1030 '~Spare MB2[32].6'; 1031 '~Spare MB2[32].7'; 1032 '~S001R13CN.I.StudWld2Rdy - Robot Stud Weld Controller 2 Not Ready MB2[32].8'; 1033 '~S001R13CN.I.Rvt2RdyToOperate - Robot Rivet Controller 2 Not Ready MB2[32].9'; 1034 '~S001R13CN.Ix.LaserWldOn - Robot Laser In No Cut MB2[32].10'; 1035 '~S001R13CN.Ix.GlassNotPres - Robot Laser Glass Not Present MB2[32].11'; 1036 '~S001R13CN.Ix.LaserHeadRdy - Robot Laser Head Not Ready MB2[32].12'; 1037 '~S001R13CN.Ix.ChillerOn - Robot Laser Chiller Not On MB2[32].13'; 1038 '~S001R13CN.Ix.GasOn - Robot Gas Not On MB2[32].14'; 1039 '~S001R13 Power Meter Not Ready MB2[32].15'; 1040 '~S001R13 No Wire Present Replace Barrel MB2[32].16'; 1041 '~S001R13 Wire Feeder Fault Timer MB2[32].17'; 1042 '~S001R13CN.Ix.NRFlt - Robot Nut Runner Not Ready MB2[32].18'; 1043 '~Spare MB2[32].19'; 1044 '~S001R13CN.M.WrongRivetAtNose - Remove Wrong Rivet At Nose MB2[32].20'; 1045 '~S001R13CN.M.DisableRbtDrvs - In Rivet Zone But Riveter Not In Auto MB2[32].21'; 1046 '~S001R13CN.I.Rvt1SystemInAuto - Rivet Controller 1 Not In Auto MB2[32].22'; 1047 '~S001R13CN.I.Rvt2SystemInAuto - Rivet Controller 2 Not In Auto MB2[32].23'; 1048 '~S001R13CN.M.RvtC1ReelCtr.DN - Reel Change Required MB2[32].24'; 1049 '~S001R13CN.M.RvtC2ReelCtr.DN - Reel Change Required MB2[32].25'; 1050 '~S001R13CN.M.AbortSkipRemain - SkipRemaining Aborted, Reset At Rbt Controller Is Required MB2[32].26'; 1051 '~Spare MB2[32].27'; 1052 '~Spare MB2[32].28'; 1053 '~Spare MB2[32].29'; 1054 '~Spare MB2[32].30'; 1055 '~Spare MB2[32].31'; 1056 '~Spare MB2[33].0'; 1057 '~Spare MB2[33].1'; 1058 '~Spare MB2[33].2'; 1059 '~Spare MB2[33].3'; 1060 '~Spare MB2[33].4'; 1061 '~Spare MB2[33].5'; 1062 '~Spare MB2[33].6'; 1063 '~Spare MB2[33].7'; 1064 '~Spare MB2[33].8'; 1065 '~Spare MB2[33].9'; 1066 '~Spare MB2[33].10'; 1067 '~Spare MB2[33].11'; 1068 '~Spare MB2[33].12'; 1069 '~Spare MB2[33].13'; 1070 '~Spare MB2[33].14'; 1071 '~Spare MB2[33].15'; 1072 '~Spare MB2[33].16'; 1073 '~Spare MB2[33].17'; 1074 '~Spare MB2[33].18'; 1075 '~Spare MB2[33].19'; 1076 '~Spare MB2[33].20'; 1077 '~Spare MB2[33].21'; 1078 '~Spare MB2[33].22'; 1079 '~Spare MB2[33].23'; 1080 '~Spare MB2[33].24'; 1081 '~Spare MB2[33].25'; 1082 '~Spare MB2[33].26'; 1083 '~Spare MB2[33].27'; 1084 '~Spare MB2[33].28'; 1085 '~Spare MB2[33].29'; 1086 '~Spare MB2[33].30'; 1087 '~Spare MB2[33].31'; 1088 '~Spare MB2[34].0'; 1089 '~Spare MB2[34].1'; 1090 '~Spare MB2[34].2'; 1091 '~Spare MB2[34].3'; 1092 '~Spare MB2[34].4'; 1093 '~Spare MB2[34].5'; 1094 '~Spare MB2[34].6'; 1095 '~Spare MB2[34].7'; 1096 '~Spare MB2[34].8'; 1097 '~Spare MB2[34].9'; 1098 '~Spare MB2[34].10'; 1099 '~Spare MB2[34].11'; 1100 '~Spare MB2[34].12'; 1101 '~Spare MB2[34].13'; 1102 '~Spare MB2[34].14'; 1103 '~Spare MB2[34].15'; 1104 '~Spare MB2[34].16'; 1105 '~Spare MB2[34].17'; 1106 '~Spare MB2[34].18'; 1107 '~Spare MB2[34].19'; 1108 '~Spare MB2[34].20'; 1109 '~Spare MB2[34].21'; 1110 '~Spare MB2[34].22'; 1111 '~Spare MB2[34].23'; 1112 '~Spare MB2[34].24'; 1113 '~Spare MB2[34].25'; 1114 '~Spare MB2[34].26'; 1115 '~Spare MB2[34].27'; 1116 '~Spare MB2[34].28'; 1117 '~Spare MB2[34].29'; 1118 '~Spare MB2[34].30'; 1119 '~Spare MB2[34].31'; 1120 '~Spare MB2[35].0'; 1121 '~Spare MB2[35].1'; 1122 '~Spare MB2[35].2'; 1123 '~Spare MB2[35].3'; 1124 '~Spare MB2[35].4'; 1125 '~Spare MB2[35].5'; 1126 '~Spare MB2[35].6'; 1127 '~Spare MB2[35].7'; 1128 '~Spare MB2[35].8'; 1129 '~Spare MB2[35].9'; 1130 '~Spare MB2[35].10'; 1131 '~Spare MB2[35].11'; 1132 '~Spare MB2[35].12'; 1133 '~Spare MB2[35].13'; 1134 '~Spare MB2[35].14'; 1135 '~Spare MB2[35].15'; 1136 '~Spare MB2[35].16'; 1137 '~Spare MB2[35].17'; 1138 '~Spare MB2[35].18'; 1139 '~Spare MB2[35].19'; 1140 '~Spare MB2[35].20'; 1141 '~Spare MB2[35].21'; 1142 '~Spare MB2[35].22'; 1143 '~Spare MB2[35].23'; 1144 '~Spare MB2[35].24'; 1145 '~Spare MB2[35].25'; 1146 '~Spare MB2[35].26'; 1147 '~Spare MB2[35].27'; 1148 '~Spare MB2[35].28'; 1149 '~Spare MB2[35].29'; 1150 '~Spare MB2[35].30'; 1151 '~Spare MB2[35].31'; 1152 '~S001R14ES1 - S001R14 EtherNet Switch Connection Inhibited MB2[36].0'; 1153 '~Spare MB2[36].1'; 1154 '~Spare MB2[36].2'; 1155 '~Spare MB2[36].3'; 1156 '~Spare MB2[36].4'; 1157 '~Spare MB2[36].5'; 1158 '~Spare MB2[36].6'; 1159 '~Spare MB2[36].7'; 1160 '~Spare MB2[36].8'; 1161 '~Spare MB2[36].9'; 1162 '~Spare MB2[36].10'; 1163 '~Spare MB2[36].11'; 1164 '~Spare MB2[36].12'; 1165 '~Spare MB2[36].13'; 1166 '~Spare MB2[36].14'; 1167 '~Spare MB2[36].15'; 1168 '~Spare MB2[36].16'; 1169 '~S001R14Sfty - Robot E-Stop Depressed MB2[36].17'; 1170 '~S001R14Sfty - Robot Safety Interface Not Enabled MB2[36].18'; 1171 '~S001R14Sfty - Robot DCS Has Been Edited MB2[36].19'; 1172 '~S001R14CN - Robot Controller Connection Inhibited MB2[36].20'; 1173 '~S001R14E#B# - Robot End Effector Module Connection Inhibited MB2[36].21'; 1174 '~S001R14E#B# - Robot End Effector Module Connection Inhibited MB2[36].22'; 1175 '~S001R14E#B# - Robot End Effector Module Connection Inhibited MB2[36].23'; 1176 '~S001R14E#B# - Robot End Effector Module Connection Inhibited MB2[36].24'; 1177 '~S001R14E#B# - Robot End Effector Module Connection Inhibited MB2[36].25'; 1178 '~S001R14E#B# - Robot End Effector Module Connection Inhibited MB2[36].26'; 1179 '~S001R14E#B# - Robot End Effector Module Connection Inhibited MB2[36].27'; 1180 '~S001R14E#B# - Robot End Effector Module Connection Inhibited MB2[36].28'; 1181 '~S001R14E#B# - Robot End Effector Module Connection Inhibited MB2[36].29'; 1182 '~Spare MB2[36].30'; 1183 '~Spare MB2[36].31'; 1184 '~Spare MB2[37].0'; 1185 '~S001R14F#B# - Robot Process I/O Connection Inhibited MB2[37].1'; 1186 '~S001R14F#B# - Robot Process I/O Connection Inhibited MB2[37].2'; 1187 '~S001R14F#B# - Robot Process I/O Connection Inhibited MB2[37].3'; 1188 '~S001R14F#B# - Robot Process I/O Connection Inhibited MB2[37].4'; 1189 '~Spare MB2[37].5'; 1190 '~Spare MB2[37].6'; 1191 '~Spare MB2[37].7'; 1192 '~Spare MB2[37].8'; 1193 '~Spare MB2[37].9'; 1194 '~S001R14CN.I.Safety - Chain Fault MB2[37].10'; 1195 '~S001R14CN.I.AirOn - Robot Air Not On MB2[37].11'; 1196 '~S001R14CN.I.RbtAuto - Robot Not in Auto MB2[37].12'; 1197 '~S001R14CN.M.InTeach - Robot In Teach MB2[37].13'; 1198 '~S001R14CN.I.AtMaintPos - Robot At Maintenace MB2[37].14'; 1199 '~S001R14CN.I.RunEnblInterruptAck - Robot In Hold MB2[37].15'; 1200 '~S001R14CN.M.MaintPosSeld - Robot Maintenance Selected MB2[37].16'; 1201 '~Spare MB2[37].17'; 1202 '~Spare MB2[37].18'; 1203 '~Spare MB2[37].19'; 1204 '~S001R14CN.I.ExtAppCommFlt - Robot Application Communication Fault MB2[37].20'; 1205 '~S001R14CN.M.AbortPickupSeld - Robot Abort Pickup Selected MB2[37].21'; 1206 '~S001R14CN.M.RetFmPounceSeld - Robot Return From Pounce Selected MB2[37].22'; 1207 '~S001R14CN.I.StudWld1 Comm Not OK MB2[37].23'; 1208 '~S001R14CN.I.StudWld2 Comm Not OK MB2[37].24'; 1209 '~S001R14CN.I.WldMode - Robot In No Weld MB2[37].25'; 1210 '~S001R14CN.I.PulledTipBypSS - Robot Pulled Tip Bypass Selected MB2[37].26'; 1211 '~S001R14CN.I.FlowNoFlowSS - Robot In No Flow MB2[37].27'; 1212 '~S001R14CN.I.RvtNoRvtSS - Robot In No Rivet MB2[37].28'; 1213 '~S001R14CN.I.WldCtrlCommOk1 - Robot Weld Controller 1 Comm Not OK MB2[37].29'; 1214 '~S001R14CN.I.WldModeStud - Robot In No Weld Stud MB2[37].30'; 1215 '~S001R14CN.Ix.MigWldNoWld - Robot In No Weld Mig MB2[37].31'; 1216 '~S001R14CN.I.StudWld1Rdy - Robot Stud Weld Controller 1 Not Ready MB2[38].0'; 1217 '~S001R14CN.I.Rvt1RdyToOperate - Robot Rivet Controller 1 Not Ready MB2[38].1'; 1218 '~S001R14CN.Ix.MigRdy - Robot Mig Weld Controller Not Ready MB2[38].2'; 1219 '~S001R14CN.Ix.MigWldNoWld - Robot In No Weld MB2[38].3'; 1220 '~Spare MB2[38].4'; 1221 '~S001R14CN.I.WldCtrlCommOk2 - Robot Weld Controller 2 Comm Not OK MB2[38].5'; 1222 '~Spare MB2[38].6'; 1223 '~Spare MB2[38].7'; 1224 '~S001R14CN.I.StudWld2Rdy - Robot Stud Weld Controller 2 Not Ready MB2[38].8'; 1225 '~S001R14CN.I.Rvt2RdyToOperate - Robot Rivet Controller 2 Not Ready MB2[38].9'; 1226 '~S001R14CN.Ix.LaserWldOn - Robot Laser In No Cut MB2[38].10'; 1227 '~S001R14CN.Ix.GlassNotPres - Robot Laser Glass Not Present MB2[38].11'; 1228 '~S001R14CN.Ix.LaserHeadRdy - Robot Laser Head Not Ready MB2[38].12'; 1229 '~S001R14CN.Ix.ChillerOn - Robot Laser Chiller Not On MB2[38].13'; 1230 '~S001R14CN.Ix.GasOn - Robot Gas Not On MB2[38].14'; 1231 '~S001R14 Power Meter Not Ready MB2[38].15'; 1232 '~S001R14 No Wire Present Replace Barrel MB2[38].16'; 1233 '~S001R14 Wire Feeder Fault Timer MB2[38].17'; 1234 '~S001R14CN.Ix.NRFlt - Robot Nut Runner Not Ready MB2[38].18'; 1235 '~Spare MB2[38].19'; 1236 '~S001R14CN.M.WrongRivetAtNose - Remove Wrong Rivet At Nose MB2[38].20'; 1237 '~S001R14CN.M.DisableRbtDrvs - In Rivet Zone But Riveter Not In Auto MB2[38].21'; 1238 '~S001R14CN.I.Rvt1SystemInAuto - Rivet Controller 1 Not In Auto MB2[38].22'; 1239 '~S001R14CN.I.Rvt2SystemInAuto - Rivet Controller 2 Not In Auto MB2[38].23'; 1240 '~S001R14CN.M.RvtC1ReelCtr.DN - Reel Change Required MB2[38].24'; 1241 '~S001R14CN.M.RvtC2ReelCtr.DN - Reel Change Required MB2[38].25'; 1242 '~S001R14CN.M.AbortSkipRemain - SkipRemaining Aborted, Reset At Rbt Controller Is Required MB2[38].26'; 1243 '~Spare MB2[38].27'; 1244 '~Spare MB2[38].28'; 1245 '~Spare MB2[38].29'; 1246 '~Spare MB2[38].30'; 1247 '~Spare MB2[38].31'; 1248 '~Spare MB2[39].0'; 1249 '~Spare MB2[39].1'; 1250 '~Spare MB2[39].2'; 1251 '~Spare MB2[39].3'; 1252 '~Spare MB2[39].4'; 1253 '~Spare MB2[39].5'; 1254 '~Spare MB2[39].6'; 1255 '~Spare MB2[39].7'; 1256 '~Spare MB2[39].8'; 1257 '~Spare MB2[39].9'; 1258 '~Spare MB2[39].10'; 1259 '~Spare MB2[39].11'; 1260 '~Spare MB2[39].12'; 1261 '~Spare MB2[39].13'; 1262 '~Spare MB2[39].14'; 1263 '~Spare MB2[39].15'; 1264 '~Spare MB2[39].16'; 1265 '~Spare MB2[39].17'; 1266 '~Spare MB2[39].18'; 1267 '~Spare MB2[39].19'; 1268 '~Spare MB2[39].20'; 1269 '~Spare MB2[39].21'; 1270 '~Spare MB2[39].22'; 1271 '~Spare MB2[39].23'; 1272 '~Spare MB2[39].24'; 1273 '~Spare MB2[39].25'; 1274 '~Spare MB2[39].26'; 1275 '~Spare MB2[39].27'; 1276 '~Spare MB2[39].28'; 1277 '~Spare MB2[39].29'; 1278 '~Spare MB2[39].30'; 1279 '~Spare MB2[39].31'; 1280 '~Spare MB2[40].0'; 1281 '~Spare MB2[40].1'; 1282 '~Spare MB2[40].2'; 1283 '~Spare MB2[40].3'; 1284 '~Spare MB2[40].4'; 1285 '~Spare MB2[40].5'; 1286 '~Spare MB2[40].6'; 1287 '~Spare MB2[40].7'; 1288 '~Spare MB2[40].8'; 1289 '~Spare MB2[40].9'; 1290 '~Spare MB2[40].10'; 1291 '~Spare MB2[40].11'; 1292 '~Spare MB2[40].12'; 1293 '~Spare MB2[40].13'; 1294 '~Spare MB2[40].14'; 1295 '~Spare MB2[40].15'; 1296 '~Spare MB2[40].16'; 1297 '~Spare MB2[40].17'; 1298 '~Spare MB2[40].18'; 1299 '~Spare MB2[40].19'; 1300 '~Spare MB2[40].20'; 1301 '~Spare MB2[40].21'; 1302 '~Spare MB2[40].22'; 1303 '~Spare MB2[40].23'; 1304 '~Spare MB2[40].24'; 1305 '~Spare MB2[40].25'; 1306 '~Spare MB2[40].26'; 1307 '~Spare MB2[40].27'; 1308 '~Spare MB2[40].28'; 1309 '~Spare MB2[40].29'; 1310 '~Spare MB2[40].30'; 1311 '~Spare MB2[40].31'; 1312 '~Spare MB2[41].0'; 1313 '~Spare MB2[41].1'; 1314 '~Spare MB2[41].2'; 1315 '~Spare MB2[41].3'; 1316 '~Spare MB2[41].4'; 1317 '~Spare MB2[41].5'; 1318 '~Spare MB2[41].6'; 1319 '~Spare MB2[41].7'; 1320 '~Spare MB2[41].8'; 1321 '~Spare MB2[41].9'; 1322 '~Spare MB2[41].10'; 1323 '~Spare MB2[41].11'; 1324 '~Spare MB2[41].12'; 1325 '~Spare MB2[41].13'; 1326 '~Spare MB2[41].14'; 1327 '~Spare MB2[41].15'; 1328 '~Spare MB2[41].16'; 1329 '~Spare MB2[41].17'; 1330 '~Spare MB2[41].18'; 1331 '~Spare MB2[41].19'; 1332 '~Spare MB2[41].20'; 1333 '~Spare MB2[41].21'; 1334 '~Spare MB2[41].22'; 1335 '~Spare MB2[41].23'; 1336 '~Spare MB2[41].24'; 1337 '~Spare MB2[41].25'; 1338 '~Spare MB2[41].26'; 1339 '~Spare MB2[41].27'; 1340 '~Spare MB2[41].28'; 1341 '~Spare MB2[41].29'; 1342 '~Spare MB2[41].30'; 1343 '~Spare MB2[41].31'; 1344 '~S001R15ES1 - S001R15 EtherNet Switch Connection Inhibited MB2[42].0'; 1345 '~Spare MB2[42].1'; 1346 '~Spare MB2[42].2'; 1347 '~Spare MB2[42].3'; 1348 '~Spare MB2[42].4'; 1349 '~Spare MB2[42].5'; 1350 '~Spare MB2[42].6'; 1351 '~Spare MB2[42].7'; 1352 '~Spare MB2[42].8'; 1353 '~Spare MB2[42].9'; 1354 '~Spare MB2[42].10'; 1355 '~Spare MB2[42].11'; 1356 '~Spare MB2[42].12'; 1357 '~Spare MB2[42].13'; 1358 '~Spare MB2[42].14'; 1359 '~Spare MB2[42].15'; 1360 '~Spare MB2[42].16'; 1361 '~S001R15Sfty - Robot E-Stop Depressed MB2[42].17'; 1362 '~S001R15Sfty - Robot Safety Interface Not Enabled MB2[42].18'; 1363 '~S001R15Sfty - Robot DCS Has Been Edited MB2[42].19'; 1364 '~S001R15CN - Robot Controller Connection Inhibited MB2[42].20'; 1365 '~S001R15E#B# - Robot End Effector Module Connection Inhibited MB2[42].21'; 1366 '~S001R15E#B# - Robot End Effector Module Connection Inhibited MB2[42].22'; 1367 '~S001R15E#B# - Robot End Effector Module Connection Inhibited MB2[42].23'; 1368 '~S001R15E#B# - Robot End Effector Module Connection Inhibited MB2[42].24'; 1369 '~S001R15E#B# - Robot End Effector Module Connection Inhibited MB2[42].25'; 1370 '~S001R15E#B# - Robot End Effector Module Connection Inhibited MB2[42].26'; 1371 '~S001R15E#B# - Robot End Effector Module Connection Inhibited MB2[42].27'; 1372 '~S001R15E#B# - Robot End Effector Module Connection Inhibited MB2[42].28'; 1373 '~S001R15E#B# - Robot End Effector Module Connection Inhibited MB2[42].29'; 1374 '~Spare MB2[42].30'; 1375 '~Spare MB2[42].31'; 1376 '~Spare MB2[43].0'; 1377 '~S001R15F#B# - Robot Process I/O Connection Inhibited MB2[43].1'; 1378 '~S001R15F#B# - Robot Process I/O Connection Inhibited MB2[43].2'; 1379 '~S001R15F#B# - Robot Process I/O Connection Inhibited MB2[43].3'; 1380 '~S001R15F#B# - Robot Process I/O Connection Inhibited MB2[43].4'; 1381 '~Spare MB2[43].5'; 1382 '~Spare MB2[43].6'; 1383 '~Spare MB2[43].7'; 1384 '~Spare MB2[43].8'; 1385 '~Spare MB2[43].9'; 1386 '~S001R15CN.I.Safety - Chain Fault MB2[43].10'; 1387 '~S001R15CN.I.AirOn - Robot Air Not On MB2[43].11'; 1388 '~S001R15CN.I.RbtAuto - Robot Not in Auto MB2[43].12'; 1389 '~S001R15CN.M.InTeach - Robot In Teach MB2[43].13'; 1390 '~S001R15CN.I.AtMaintPos - Robot At Maintenace MB2[43].14'; 1391 '~S001R15CN.I.RunEnblInterruptAck - Robot In Hold MB2[43].15'; 1392 '~S001R15CN.M.MaintPosSeld - Robot Maintenance Selected MB2[43].16'; 1393 '~Spare MB2[43].17'; 1394 '~Spare MB2[43].18'; 1395 '~Spare MB2[43].19'; 1396 '~S001R15CN.I.ExtAppCommFlt - Robot Application Communication Fault MB2[43].20'; 1397 '~S001R15CN.M.AbortPickupSeld - Robot Abort Pickup Selected MB2[43].21'; 1398 '~S001R15CN.M.RetFmPounceSeld - Robot Return From Pounce Selected MB2[43].22'; 1399 '~S001R15CN.I.StudWld1 Comm Not OK MB2[43].23'; 1400 '~S001R15CN.I.StudWld2 Comm Not OK MB2[43].24'; 1401 '~S001R15CN.I.WldMode - Robot In No Weld MB2[43].25'; 1402 '~S001R15CN.I.PulledTipBypSS - Robot Pulled Tip Bypass Selected MB2[43].26'; 1403 '~S001R15CN.I.FlowNoFlowSS - Robot In No Flow MB2[43].27'; 1404 '~S001R15CN.I.RvtNoRvtSS - Robot In No Rivet MB2[43].28'; 1405 '~S001R15CN.I.WldCtrlCommOk1 - Robot Weld Controller 1 Comm Not OK MB2[43].29'; 1406 '~S001R15CN.I.WldModeStud - Robot In No Weld Stud MB2[43].30'; 1407 '~S001R15CN.Ix.MigWldNoWld - Robot In No Weld Mig MB2[43].31'; 1408 '~S001R15CN.I.StudWld1Rdy - Robot Stud Weld Controller 1 Not Ready MB2[44].0'; 1409 '~S001R15CN.I.Rvt1RdyToOperate - Robot Rivet Controller 1 Not Ready MB2[44].1'; 1410 '~S001R15CN.Ix.MigRdy - Robot Mig Weld Controller Not Ready MB2[44].2'; 1411 '~S001R15CN.Ix.MigWldNoWld - Robot In No Weld MB2[44].3'; 1412 '~Spare MB2[44].4'; 1413 '~S001R15CN.I.WldCtrlCommOk2 - Robot Weld Controller 2 Comm Not OK MB2[44].5'; 1414 '~Spare MB2[44].6'; 1415 '~Spare MB2[44].7'; 1416 '~S001R15CN.I.StudWld2Rdy - Robot Stud Weld Controller 2 Not Ready MB2[44].8'; 1417 '~S001R15CN.I.Rvt2RdyToOperate - Robot Rivet Controller 2 Not Ready MB2[44].9'; 1418 '~S001R15CN.Ix.LaserWldOn - Robot Laser In No Cut MB2[44].10'; 1419 '~S001R15CN.Ix.GlassNotPres - Robot Laser Glass Not Present MB2[44].11'; 1420 '~S001R15CN.Ix.LaserHeadRdy - Robot Laser Head Not Ready MB2[44].12'; 1421 '~S001R15CN.Ix.ChillerOn - Robot Laser Chiller Not On MB2[44].13'; 1422 '~S001R15CN.Ix.GasOn - Robot Gas Not On MB2[44].14'; 1423 '~S001R15 Power Meter Not Ready MB2[44].15'; 1424 '~S001R15 No Wire Present Replace Barrel MB2[44].16'; 1425 '~S001R15 Wire Feeder Fault Timer MB2[44].17'; 1426 '~S001R15CN.Ix.NRFlt - Robot Nut Runner Not Ready MB2[44].18'; 1427 '~Spare MB2[44].19'; 1428 '~S001R15CN.M.WrongRivetAtNose - Remove Wrong Rivet At Nose MB2[44].20'; 1429 '~S001R15CN.M.DisableRbtDrvs - In Rivet Zone But Riveter Not In Auto MB2[44].21'; 1430 '~S001R15CN.I.Rvt1SystemInAuto - Rivet Controller 1 Not In Auto MB2[44].22'; 1431 '~S001R15CN.I.Rvt2SystemInAuto - Rivet Controller 2 Not In Auto MB2[44].23'; 1432 '~S001R15CN.M.RvtC1ReelCtr.DN - Reel Change Required MB2[44].24'; 1433 '~S001R15CN.M.RvtC2ReelCtr.DN - Reel Change Required MB2[44].25'; 1434 '~S001R15CN.M.AbortSkipRemain - SkipRemaining Aborted, Reset At Rbt Controller Is Required MB2[44].26'; 1435 '~Spare MB2[44].27'; 1436 '~Spare MB2[44].28'; 1437 '~Spare MB2[44].29'; 1438 '~Spare MB2[44].30'; 1439 '~Spare MB2[44].31'; 1440 '~Spare MB2[45].0'; 1441 '~Spare MB2[45].1'; 1442 '~Spare MB2[45].2'; 1443 '~Spare MB2[45].3'; 1444 '~Spare MB2[45].4'; 1445 '~Spare MB2[45].5'; 1446 '~Spare MB2[45].6'; 1447 '~Spare MB2[45].7'; 1448 '~Spare MB2[45].8'; 1449 '~Spare MB2[45].9'; 1450 '~Spare MB2[45].10'; 1451 '~Spare MB2[45].11'; 1452 '~Spare MB2[45].12'; 1453 '~Spare MB2[45].13'; 1454 '~Spare MB2[45].14'; 1455 '~Spare MB2[45].15'; 1456 '~Spare MB2[45].16'; 1457 '~Spare MB2[45].17'; 1458 '~Spare MB2[45].18'; 1459 '~Spare MB2[45].19'; 1460 '~Spare MB2[45].20'; 1461 '~Spare MB2[45].21'; 1462 '~Spare MB2[45].22'; 1463 '~Spare MB2[45].23'; 1464 '~Spare MB2[45].24'; 1465 '~Spare MB2[45].25'; 1466 '~Spare MB2[45].26'; 1467 '~Spare MB2[45].27'; 1468 '~Spare MB2[45].28'; 1469 '~Spare MB2[45].29'; 1470 '~Spare MB2[45].30'; 1471 '~Spare MB2[45].31'; 1472 '~Spare MB2[46].0'; 1473 '~Spare MB2[46].1'; 1474 '~Spare MB2[46].2'; 1475 '~Spare MB2[46].3'; 1476 '~Spare MB2[46].4'; 1477 '~Spare MB2[46].5'; 1478 '~Spare MB2[46].6'; 1479 '~Spare MB2[46].7'; 1480 '~Spare MB2[46].8'; 1481 '~Spare MB2[46].9'; 1482 '~Spare MB2[46].10'; 1483 '~Spare MB2[46].11'; 1484 '~Spare MB2[46].12'; 1485 '~Spare MB2[46].13'; 1486 '~Spare MB2[46].14'; 1487 '~Spare MB2[46].15'; 1488 '~Spare MB2[46].16'; 1489 '~Spare MB2[46].17'; 1490 '~Spare MB2[46].18'; 1491 '~Spare MB2[46].19'; 1492 '~Spare MB2[46].20'; 1493 '~Spare MB2[46].21'; 1494 '~Spare MB2[46].22'; 1495 '~Spare MB2[46].23'; 1496 '~Spare MB2[46].24'; 1497 '~Spare MB2[46].25'; 1498 '~Spare MB2[46].26'; 1499 '~Spare MB2[46].27'; 1500 '~Spare MB2[46].28'; 1501 '~Spare MB2[46].29'; 1502 '~Spare MB2[46].30'; 1503 '~Spare MB2[46].31'; 1504 '~Spare MB2[47].0'; 1505 '~Spare MB2[47].1'; 1506 '~Spare MB2[47].2'; 1507 '~Spare MB2[47].3'; 1508 '~Spare MB2[47].4'; 1509 '~Spare MB2[47].5'; 1510 '~Spare MB2[47].6'; 1511 '~Spare MB2[47].7'; 1512 '~Spare MB2[47].8'; 1513 '~Spare MB2[47].9'; 1514 '~Spare MB2[47].10'; 1515 '~Spare MB2[47].11'; 1516 '~Spare MB2[47].12'; 1517 '~Spare MB2[47].13'; 1518 '~Spare MB2[47].14'; 1519 '~Spare MB2[47].15'; 1520 '~Spare MB2[47].16'; 1521 '~Spare MB2[47].17'; 1522 '~Spare MB2[47].18'; 1523 '~Spare MB2[47].19'; 1524 '~Spare MB2[47].20'; 1525 '~Spare MB2[47].21'; 1526 '~Spare MB2[47].22'; 1527 '~Spare MB2[47].23'; 1528 '~Spare MB2[47].24'; 1529 '~Spare MB2[47].25'; 1530 '~Spare MB2[47].26'; 1531 '~Spare MB2[47].27'; 1532 '~Spare MB2[47].28'; 1533 '~Spare MB2[47].29'; 1534 '~Spare MB2[47].30'; 1535 '~Spare MB2[47].31'; 1536 '~S001R16ES1 - S001R16 EtherNet Switch Connection Inhibited MB2[48].0'; 1537 '~Spare MB2[48].1'; 1538 '~Spare MB2[48].2'; 1539 '~Spare MB2[48].3'; 1540 '~Spare MB2[48].4'; 1541 '~Spare MB2[48].5'; 1542 '~Spare MB2[48].6'; 1543 '~Spare MB2[48].7'; 1544 '~Spare MB2[48].8'; 1545 '~Spare MB2[48].9'; 1546 '~Spare MB2[48].10'; 1547 '~Spare MB2[48].11'; 1548 '~Spare MB2[48].12'; 1549 '~Spare MB2[48].13'; 1550 '~Spare MB2[48].14'; 1551 '~Spare MB2[48].15'; 1552 '~Spare MB2[48].16'; 1553 '~S001R16Sfty - Robot E-Stop Depressed MB2[48].17'; 1554 '~S001R16Sfty - Robot Safety Interface Not Enabled MB2[48].18'; 1555 '~S001R16Sfty - Robot DCS Has Been Edited MB2[48].19'; 1556 '~S001R16CN - Robot Controller Connection Inhibited MB2[48].20'; 1557 '~S001R16E#B# - Robot End Effector Module Connection Inhibited MB2[48].21'; 1558 '~S001R16E#B# - Robot End Effector Module Connection Inhibited MB2[48].22'; 1559 '~S001R16E#B# - Robot End Effector Module Connection Inhibited MB2[48].23'; 1560 '~S001R16E#B# - Robot End Effector Module Connection Inhibited MB2[48].24'; 1561 '~S001R16E#B# - Robot End Effector Module Connection Inhibited MB2[48].25'; 1562 '~S001R16E#B# - Robot End Effector Module Connection Inhibited MB2[48].26'; 1563 '~S001R16E#B# - Robot End Effector Module Connection Inhibited MB2[48].27'; 1564 '~S001R16E#B# - Robot End Effector Module Connection Inhibited MB2[48].28'; 1565 '~S001R16E#B# - Robot End Effector Module Connection Inhibited MB2[48].29'; 1566 '~Spare MB2[48].30'; 1567 '~Spare MB2[48].31'; 1568 '~Spare MB2[49].0'; 1569 '~S001R16F#B# - Robot Process I/O Connection Inhibited MB2[49].1'; 1570 '~S001R16F#B# - Robot Process I/O Connection Inhibited MB2[49].2'; 1571 '~S001R16F#B# - Robot Process I/O Connection Inhibited MB2[49].3'; 1572 '~S001R16F#B# - Robot Process I/O Connection Inhibited MB2[49].4'; 1573 '~Spare MB2[49].5'; 1574 '~Spare MB2[49].6'; 1575 '~Spare MB2[49].7'; 1576 '~Spare MB2[49].8'; 1577 '~Spare MB2[49].9'; 1578 '~S001R16CN.I.Safety - Chain Fault MB2[49].10'; 1579 '~S001R16CN.I.AirOn - Robot Air Not On MB2[49].11'; 1580 '~S001R16CN.I.RbtAuto - Robot Not in Auto MB2[49].12'; 1581 '~S001R16CN.M.InTeach - Robot In Teach MB2[49].13'; 1582 '~S001R16CN.I.AtMaintPos - Robot At Maintenace MB2[49].14'; 1583 '~S001R16CN.I.RunEnblInterruptAck - Robot In Hold MB2[49].15'; 1584 '~S001R16CN.M.MaintPosSeld - Robot Maintenance Selected MB2[49].16'; 1585 '~Spare MB2[49].17'; 1586 '~Spare MB2[49].18'; 1587 '~Spare MB2[49].19'; 1588 '~S001R16CN.I.ExtAppCommFlt - Robot Application Communication Fault MB2[49].20'; 1589 '~S001R16CN.M.AbortPickupSeld - Robot Abort Pickup Selected MB2[49].21'; 1590 '~S001R16CN.M.RetFmPounceSeld - Robot Return From Pounce Selected MB2[49].22'; 1591 '~S001R16CN.I.StudWld1 Comm Not OK MB2[49].23'; 1592 '~S001R16CN.I.StudWld2 Comm Not OK MB2[49].24'; 1593 '~S001R16CN.I.WldMode - Robot In No Weld MB2[49].25'; 1594 '~S001R16CN.I.PulledTipBypSS - Robot Pulled Tip Bypass Selected MB2[49].26'; 1595 '~S001R16CN.I.FlowNoFlowSS - Robot In No Flow MB2[49].27'; 1596 '~S001R16CN.I.RvtNoRvtSS - Robot In No Rivet MB2[49].28'; 1597 '~S001R16CN.I.WldCtrlCommOk1 - Robot Weld Controller 1 Comm Not OK MB2[49].29'; 1598 '~S001R16CN.I.WldModeStud - Robot In No Weld Stud MB2[49].30'; 1599 '~S001R16CN.Ix.MigWldNoWld - Robot In No Weld Mig MB2[49].31'; 1600 '~S001R16CN.I.StudWld1Rdy - Robot Stud Weld Controller 1 Not Ready MB2[50].0'; 1601 '~S001R16CN.I.Rvt1RdyToOperate - Robot Rivet Controller 1 Not Ready MB2[50].1'; 1602 '~S001R16CN.Ix.MigRdy - Robot Mig Weld Controller Not Ready MB2[50].2'; 1603 '~S001R16CN.Ix.MigWldNoWld - Robot In No Weld MB2[50].3'; 1604 '~Spare MB2[50].4'; 1605 '~S001R16CN.I.WldCtrlCommOk2 - Robot Weld Controller 2 Comm Not OK MB2[50].5'; 1606 '~Spare MB2[50].6'; 1607 '~Spare MB2[50].7'; 1608 '~S001R16CN.I.StudWld2Rdy - Robot Stud Weld Controller 2 Not Ready MB2[50].8'; 1609 '~S001R16CN.I.Rvt2RdyToOperate - Robot Rivet Controller 2 Not Ready MB2[50].9'; 1610 '~S001R16CN.Ix.LaserWldOn - Robot Laser In No Cut MB2[50].10'; 1611 '~S001R16CN.Ix.GlassNotPres - Robot Laser Glass Not Present MB2[50].11'; 1612 '~S001R16CN.Ix.LaserHeadRdy - Robot Laser Head Not Ready MB2[50].12'; 1613 '~S001R16CN.Ix.ChillerOn - Robot Laser Chiller Not On MB2[50].13'; 1614 '~S001R16CN.Ix.GasOn - Robot Gas Not On MB2[50].14'; 1615 '~S001R16 Power Meter Not Ready MB2[50].15'; 1616 '~S001R16 No Wire Present Replace Barrel MB2[50].16'; 1617 '~S001R16 Wire Feeder Fault Timer MB2[50].17'; 1618 '~S001R16CN.Ix.NRFlt - Robot Nut Runner Not Ready MB2[50].18'; 1619 '~Spare MB2[50].19'; 1620 '~S001R16CN.M.WrongRivetAtNose - Remove Wrong Rivet At Nose MB2[50].20'; 1621 '~S001R16CN.M.DisableRbtDrvs - In Rivet Zone But Riveter Not In Auto MB2[50].21'; 1622 '~S001R16CN.I.Rvt1SystemInAuto - Rivet Controller 1 Not In Auto MB2[50].22'; 1623 '~S001R16CN.I.Rvt2SystemInAuto - Rivet Controller 2 Not In Auto MB2[50].23'; 1624 '~S001R16CN.M.RvtC1ReelCtr.DN - Reel Change Required MB2[50].24'; 1625 '~S001R16CN.M.RvtC2ReelCtr.DN - Reel Change Required MB2[50].25'; 1626 '~S001R16CN.M.AbortSkipRemain - SkipRemaining Aborted, Reset At Rbt Controller Is Required MB2[50].26'; 1627 '~Spare MB2[50].27'; 1628 '~Spare MB2[50].28'; 1629 '~Spare MB2[50].29'; 1630 '~Spare MB2[50].30'; 1631 '~Spare MB2[50].31'; 1632 '~Spare MB2[51].0'; 1633 '~Spare MB2[51].1'; 1634 '~Spare MB2[51].2'; 1635 '~Spare MB2[51].3'; 1636 '~Spare MB2[51].4'; 1637 '~Spare MB2[51].5'; 1638 '~Spare MB2[51].6'; 1639 '~Spare MB2[51].7'; 1640 '~Spare MB2[51].8'; 1641 '~Spare MB2[51].9'; 1642 '~Spare MB2[51].10'; 1643 '~Spare MB2[51].11'; 1644 '~Spare MB2[51].12'; 1645 '~Spare MB2[51].13'; 1646 '~Spare MB2[51].14'; 1647 '~Spare MB2[51].15'; 1648 '~Spare MB2[51].16'; 1649 '~Spare MB2[51].17'; 1650 '~Spare MB2[51].18'; 1651 '~Spare MB2[51].19'; 1652 '~Spare MB2[51].20'; 1653 '~Spare MB2[51].21'; 1654 '~Spare MB2[51].22'; 1655 '~Spare MB2[51].23'; 1656 '~Spare MB2[51].24'; 1657 '~Spare MB2[51].25'; 1658 '~Spare MB2[51].26'; 1659 '~Spare MB2[51].27'; 1660 '~Spare MB2[51].28'; 1661 '~Spare MB2[51].29'; 1662 '~Spare MB2[51].30'; 1663 '~Spare MB2[51].31'; 1664 '~Spare MB2[52].0'; 1665 '~Spare MB2[52].1'; 1666 '~Spare MB2[52].2'; 1667 '~Spare MB2[52].3'; 1668 '~Spare MB2[52].4'; 1669 '~Spare MB2[52].5'; 1670 '~Spare MB2[52].6'; 1671 '~Spare MB2[52].7'; 1672 '~Spare MB2[52].8'; 1673 '~Spare MB2[52].9'; 1674 '~Spare MB2[52].10'; 1675 '~Spare MB2[52].11'; 1676 '~Spare MB2[52].12'; 1677 '~Spare MB2[52].13'; 1678 '~Spare MB2[52].14'; 1679 '~Spare MB2[52].15'; 1680 '~Spare MB2[52].16'; 1681 '~Spare MB2[52].17'; 1682 '~Spare MB2[52].18'; 1683 '~Spare MB2[52].19'; 1684 '~Spare MB2[52].20'; 1685 '~Spare MB2[52].21'; 1686 '~Spare MB2[52].22'; 1687 '~Spare MB2[52].23'; 1688 '~Spare MB2[52].24'; 1689 '~Spare MB2[52].25'; 1690 '~Spare MB2[52].26'; 1691 '~Spare MB2[52].27'; 1692 '~Spare MB2[52].28'; 1693 '~Spare MB2[52].29'; 1694 '~Spare MB2[52].30'; 1695 '~Spare MB2[52].31'; 1696 '~Spare MB2[53].0'; 1697 '~Spare MB2[53].1'; 1698 '~Spare MB2[53].2'; 1699 '~Spare MB2[53].3'; 1700 '~Spare MB2[53].4'; 1701 '~Spare MB2[53].5'; 1702 '~Spare MB2[53].6'; 1703 '~Spare MB2[53].7'; 1704 '~Spare MB2[53].8'; 1705 '~Spare MB2[53].9'; 1706 '~Spare MB2[53].10'; 1707 '~Spare MB2[53].11'; 1708 '~Spare MB2[53].12'; 1709 '~Spare MB2[53].13'; 1710 '~Spare MB2[53].14'; 1711 '~Spare MB2[53].15'; 1712 '~Spare MB2[53].16'; 1713 '~Spare MB2[53].17'; 1714 '~Spare MB2[53].18'; 1715 '~Spare MB2[53].19'; 1716 '~Spare MB2[53].20'; 1717 '~Spare MB2[53].21'; 1718 '~Spare MB2[53].22'; 1719 '~Spare MB2[53].23'; 1720 '~Spare MB2[53].24'; 1721 '~Spare MB2[53].25'; 1722 '~Spare MB2[53].26'; 1723 '~Spare MB2[53].27'; 1724 '~Spare MB2[53].28'; 1725 '~Spare MB2[53].29'; 1726 '~Spare MB2[53].30'; 1727 '~Spare MB2[53].31'; 1728 '~Spare MB2[54].0'; 1729 '~Spare MB2[54].1'; 1730 '~Spare MB2[54].2'; 1731 '~Spare MB2[54].3'; 1732 '~Spare MB2[54].4'; 1733 '~Spare MB2[54].5'; 1734 '~Spare MB2[54].6'; 1735 '~Spare MB2[54].7'; 1736 '~Spare MB2[54].8'; 1737 '~Spare MB2[54].9'; 1738 '~Spare MB2[54].10'; 1739 '~Spare MB2[54].11'; 1740 '~Spare MB2[54].12'; 1741 '~Spare MB2[54].13'; 1742 '~Spare MB2[54].14'; 1743 '~Spare MB2[54].15'; 1744 '~Spare MB2[54].16'; 1745 '~Spare MB2[54].17'; 1746 '~Spare MB2[54].18'; 1747 '~Spare MB2[54].19'; 1748 '~Spare MB2[54].20'; 1749 '~Spare MB2[54].21'; 1750 '~Spare MB2[54].22'; 1751 '~Spare MB2[54].23'; 1752 '~Spare MB2[54].24'; 1753 '~Spare MB2[54].25'; 1754 '~Spare MB2[54].26'; 1755 '~Spare MB2[54].27'; 1756 '~Spare MB2[54].28'; 1757 '~Spare MB2[54].29'; 1758 '~Spare MB2[54].30'; 1759 '~Spare MB2[54].31'; 1760 '~Spare MB2[55].0'; 1761 '~Spare MB2[55].1'; 1762 '~Spare MB2[55].2'; 1763 '~Spare MB2[55].3'; 1764 '~Spare MB2[55].4'; 1765 '~Spare MB2[55].5'; 1766 '~Spare MB2[55].6'; 1767 '~Spare MB2[55].7'; 1768 '~Spare MB2[55].8'; 1769 '~Spare MB2[55].9'; 1770 '~Spare MB2[55].10'; 1771 '~Spare MB2[55].11'; 1772 '~Spare MB2[55].12'; 1773 '~Spare MB2[55].13'; 1774 '~Spare MB2[55].14'; 1775 '~Spare MB2[55].15'; 1776 '~Spare MB2[55].16'; 1777 '~Spare MB2[55].17'; 1778 '~Spare MB2[55].18'; 1779 '~Spare MB2[55].19'; 1780 '~Spare MB2[55].20'; 1781 '~Spare MB2[55].21'; 1782 '~Spare MB2[55].22'; 1783 '~Spare MB2[55].23'; 1784 '~Spare MB2[55].24'; 1785 '~Spare MB2[55].25'; 1786 '~Spare MB2[55].26'; 1787 '~Spare MB2[55].27'; 1788 '~Spare MB2[55].28'; 1789 '~Spare MB2[55].29'; 1790 '~Spare MB2[55].30'; 1791 '~Spare MB2[55].31'; 1792 '~Spare MB2[56].0'; 1793 '~Spare MB2[56].1'; 1794 '~S002LS1Sfty - Operator 1 E-Stop Depressed MB2[56].2'; 1795 '~S002LS1Sfty - Operator 2 E-Stop Depressed MB2[56].3'; 1796 '~Spare MB2[56].4'; 1797 '~Spare MB2[56].5'; 1798 '~Spare MB2[56].6'; 1799 '~Spare MB2[56].7'; 1800 '~Spare MB2[56].8'; 1801 '~Spare MB2[56].9'; 1802 '~S002LS1Sfty - Line Access Light Screen Faulted MB2[56].10'; 1803 '~S002LS1Sfty - Operator 1 Light Screen Faulted MB2[56].11'; 1804 '~S002LS1Sfty - Operator 2 Light Screen Faulted MB2[56].12'; 1805 '~S002LS1Sfty - Operator 3 Light Screen Faulted MB2[56].13'; 1806 '~Spare MB2[56].14'; 1807 '~Spare MB2[56].15'; 1808 '~Spare MB2[56].16'; 1809 '~Spare MB2[56].17'; 1810 '~S002LS2Sfty - Operator 1 E-Stop Depressed MB2[56].18'; 1811 '~S002LS2Sfty - Operator 2 E-Stop Depressed MB2[56].19'; 1812 '~Spare MB2[56].20'; 1813 '~Spare MB2[56].21'; 1814 '~Spare MB2[56].22'; 1815 '~Spare MB2[56].23'; 1816 '~Spare MB2[56].24'; 1817 '~Spare MB2[56].25'; 1818 '~S002LS2Sfty - Line Access Light Screen Faulted MB2[56].26'; 1819 '~S002LS2Sfty - Operator 1 Light Screen Faulted MB2[56].27'; 1820 '~S002LS2Sfty - Operator 2 Light Screen Faulted MB2[56].28'; 1821 '~S002LS2Sfty - Operator 3 Light Screen Faulted MB2[56].29'; 1822 '~Spare MB2[56].30'; 1823 '~Spare MB2[56].31'; 1824 '~S002TT1DES1 - S002TT1 EtherNet Switch Connection Inhibited MB2[57].0'; 1825 '~Spare MB2[57].1'; 1826 '~Spare MB2[57].2'; 1827 '~S002TT1DES2 - S002TT1 EtherNet Switch Connection Inhibited MB2[57].3'; 1828 '~Spare MB2[57].4'; 1829 '~Spare MB2[57].5'; 1830 '~Spare MB2[57].6'; 1831 '~Spare MB2[57].7'; 1832 '~Spare MB2[57].8'; 1833 '~Spare MB2[57].9'; 1834 '~Spare MB2[57].10'; 1835 '~S002TT1.M.SafetySwOk - Turn Table Drive Pnl Disconnect Not On MB2[57].11'; 1836 '~S002TT1.M.SftyPinsOk - Turn Table Safety Pins Not In Storage MB2[57].12'; 1837 '~S002TT1.M.AirOn - Turn Table Air Pressure Not Ok MB2[57].13'; 1838 '~S002TT1 - Turn Table Safety Pin 1 Not In Storage MB2[57].14'; 1839 '~S002TT1DSfty- Turn Table Safety Contactor #1 Still On MB2[57].15'; 1840 '~S002TT1DSfty- Turn Table Safety Contactor #2 Still On MB2[57].16'; 1841 '~Spare MB2[57].17'; 1842 '~Spare MB2[57].18'; 1843 '~Spare MB2[57].19'; 1844 '~S002TT1DSfty- Turn Table Motor Brake Contactor #1 BRCR1 Still On MB2[57].20'; 1845 '~S002TT1DSfty- Turn Table Motor Brake Contactor #1 BRCR1 Not On MB2[57].21'; 1846 '~S002TT1DSfty- Turn Table Motor Brake Contactor #2 BRCR2 Still On MB2[57].22'; 1847 '~S002TT1DSfty- Turn Table Motor Brake Contactor #2 BRCR2 Not On MB2[57].23'; 1848 '~Spare MB2[57].24'; 1849 '~Spare MB2[57].25'; 1850 '~Spare MB2[57].26'; 1851 '~S002TT1DV1 - VFD Connection Inhibited MB2[57].27'; 1852 '~Spare MB2[57].28'; 1853 '~Spare MB2[57].29'; 1854 '~Spare MB2[57].30'; 1855 '~Spare MB2[57].31'; 1856 '~Spare MB2[58].0'; 1857 '~Spare MB2[58].1'; 1858 '~Spare MB2[58].2'; 1859 '~Spare MB2[58].3'; 1860 '~Spare MB2[58].4'; 1861 '~Spare MB2[58].5'; 1862 '~Spare MB2[58].6'; 1863 '~Spare MB2[58].7'; 1864 '~Spare MB2[58].8'; 1865 '~Spare MB2[58].9'; 1866 '~Spare MB2[58].10'; 1867 '~Spare MB2[58].11'; 1868 '~Spare MB2[58].12'; 1869 '~Spare MB2[58].13'; 1870 '~Spare MB2[58].14'; 1871 '~Spare MB2[58].15'; 1872 '~Spare MB2[58].16'; 1873 '~Spare MB2[58].17'; 1874 '~Spare MB2[58].18'; 1875 '~Spare MB2[58].19'; 1876 '~Spare MB2[58].20'; 1877 '~Spare MB2[58].21'; 1878 '~Spare MB2[58].22'; 1879 '~Spare MB2[58].23'; 1880 '~Spare MB2[58].24'; 1881 '~Spare MB2[58].25'; 1882 '~Spare MB2[58].26'; 1883 '~Spare MB2[58].27'; 1884 '~Spare MB2[58].28'; 1885 '~Spare MB2[58].29'; 1886 '~Spare MB2[58].30'; 1887 '~Spare MB2[58].31'; 1888 '~S001_002PRBDES1 - S001_002PRB EtherNet Switch Connection Inhibited MB2[59].0'; 1889 '~Spare MB2[59].1'; 1890 '~Spare MB2[59].2'; 1891 '~S001_002PRBDV1 - Module Connection Inhibited MB2[59].3'; 1892 '~S001_002PRBDC - Module Connection Inhibited MB2[59].4'; 1893 '~S001_002PRB1B1 - Module Connection Inhibited MB2[59].5'; 1894 '~S001_002PRB1B2 - Module Connection Inhibited MB2[59].6'; 1895 '~S001_002PRBDV2 - Module Connection Inhibited MB2[59].7'; 1896 '~S001_002PRB Panel Disconnect Off MB2[59].8'; 1897 '~Spare MB2[59].9'; 1898 '~Spare MB2[59].10'; 1899 '~Spare MB2[59].11'; 1900 '~Spare MB2[59].12'; 1901 '~S001PRB In Station Pallet/Skid Hold MB2[59].13'; 1902 '~S002PRB In Station Pallet/Skid Hold MB2[59].14'; 1903 '~Spare MB2[59].15'; 1904 '~Spare MB2[59].16'; 1905 '~Spare MB2[59].17'; 1906 '~Spare MB2[59].18'; 1907 '~Spare MB2[59].19'; 1908 '~Spare MB2[59].20'; 1909 '~Spare MB2[59].21'; 1910 '~Spare MB2[59].22'; 1911 '~Spare MB2[59].23'; 1912 '~Spare MB2[59].24'; 1913 '~Spare MB2[59].25'; 1914 '~Spare MB2[59].26'; 1915 '~Spare MB2[59].27'; 1916 '~Spare MB2[59].28'; 1917 '~Spare MB2[59].29'; 1918 '~Spare MB2[59].30'; 1919 '~S002LFT Lifter Safety Pin Fault MB2[59].31'; 1920 '~S003TL1DES1 - S003TL1 EtherNet Switch Connection Inhibited MB2[60].0'; 1921 '~Spare MB2[60].1'; 1922 '~Spare MB2[60].2'; 1923 '~Spare MB2[60].3'; 1924 '~Spare MB2[60].4'; 1925 '~Spare MB2[60].5'; 1926 '~Spare MB2[60].6'; 1927 '~Spare MB2[60].7'; 1928 '~Spare MB2[60].8'; 1929 '~Spare MB2[60].9'; 1930 '~Spare MB2[60].10'; 1931 '~S003TL1.M.SafetySwOk - Tool-Tray Drive Pnl Safety Switch Not On MB2[60].11'; 1932 '~S003TL1.M.SftyPinsOk - Tool-Tray Safety Pin Not In Storage MB2[60].12'; 1933 '~S003TL1.M.AirOn - Tool-Tray Air Pressure Not Ok MB2[60].13'; 1934 '~S003TL1 - Tool-Tray Safety Pin 1 Not In Storage MB2[60].14'; 1935 '~Spare MB2[60].15'; 1936 '~Spare MB2[60].16'; 1937 '~Spare MB2[60].17'; 1938 '~Spare MB2[60].18'; 1939 '~Spare MB2[60].19'; 1940 '~Spare MB2[60].20'; 1941 '~Spare MB2[60].21'; 1942 '~Spare MB2[60].22'; 1943 '~Spare MB2[60].23'; 1944 '~Spare MB2[60].24'; 1945 '~Spare MB2[60].25'; 1946 '~Spare MB2[60].26'; 1947 '~S003TL1DV1 - VFD Connection Inhibited MB2[60].27'; 1948 '~Spare MB2[60].28'; 1949 '~Spare MB2[60].29'; 1950 '~Spare MB2[60].30'; 1951 '~Spare MB2[60].31'; 1952 '~S002CV1DES1 - S002CV1 EtherNet Switch Connection Inhibited MB2[61].0'; 1953 '~Spare MB2[61].1'; 1954 '~Spare MB2[61].2'; 1955 '~Spare MB2[61].3'; 1956 '~Spare MB2[61].4'; 1957 '~Spare MB2[61].5'; 1958 '~Spare MB2[61].6'; 1959 '~Spare MB2[61].7'; 1960 '~Spare MB2[61].8'; 1961 '~Spare MB2[61].9'; 1962 '~Spare MB2[61].10'; 1963 '~S002CV1 - Conveyor Panel Safety Switch Not On MB2[61].11'; 1964 '~Spare MB2[61].12'; 1965 '~Spare MB2[61].13'; 1966 '~S002CV1Sfty- Conveyor Safety Contactor #1 Still On MB2[61].14'; 1967 '~S002CV1Sfty- Conveyor Safety Contactor #1 Not On MB2[61].15'; 1968 '~Spare MB2[61].16'; 1969 '~Spare MB2[61].17'; 1970 '~Spare MB2[61].18'; 1971 '~Spare MB2[61].19'; 1972 '~Spare MB2[61].20'; 1973 '~Spare MB2[61].21'; 1974 '~Spare MB2[61].22'; 1975 '~Spare MB2[61].23'; 1976 '~S002CV1DB1 - Module Connection Inhibited MB2[61].24'; 1977 '~Spare MB2[61].25'; 1978 '~Spare MB2[61].26'; 1979 '~Spare MB2[61].27'; 1980 '~S002CV1DC - Conveyor Drive Point I/O Connection Inhibited MB2[61].28'; 1981 '~Spare MB2[61].29'; 1982 '~Spare MB2[61].30'; 1983 '~Spare MB2[61].31'; 1984 '~Spare MB2[62].0'; 1985 '~Spare MB2[62].1'; 1986 '~Spare MB2[62].2'; 1987 '~Spare MB2[62].3'; 1988 '~S002CV1Sfty - Conveyor Start / Stop PB Depressed MB2[62].4'; 1989 '~Spare MB2[62].5'; 1990 '~Spare MB2[62].6'; 1991 '~Spare MB2[62].7'; 1992 '~Spare MB2[62].8'; 1993 '~Spare MB2[62].9'; 1994 '~Spare MB2[62].10'; 1995 '~Spare MB2[62].11'; 1996 '~Spare MB2[62].12'; 1997 '~Spare MB2[62].13'; 1998 '~Spare MB2[62].14'; 1999 '~Spare MB2[62].15'; 2000 '~Spare MB2[62].16'; 2001 '~Spare MB2[62].17'; 2002 '~Spare MB2[62].18'; 2003 '~Spare MB2[62].19'; 2004 '~Spare MB2[62].20'; 2005 '~Spare MB2[62].21'; 2006 '~Spare MB2[62].22'; 2007 '~Spare MB2[62].23'; 2008 '~Spare MB2[62].24'; 2009 '~Spare MB2[62].25'; 2010 '~Spare MB2[62].26'; 2011 '~Spare MB2[62].27'; 2012 '~Spare MB2[62].28'; 2013 '~Spare MB2[62].29'; 2014 '~Spare MB2[62].30'; 2015 '~Spare MB2[62].31'; 2016 '~S001CV1DES1 - S001CV1 EtherNet Switch Connection Inhibited MB2[63].0'; 2017 '~Spare MB2[63].1'; 2018 '~Spare MB2[63].2'; 2019 '~S001CV1DC - Drive I/O Connection Inhibited MB2[63].3'; 2020 '~S001CV1B1 - Module Connection Inhibited MB2[63].4'; 2021 '~Spare MB2[63].5'; 2022 '~Spare MB2[63].6'; 2023 '~Spare MB2[63].7'; 2024 '~Spare MB2[63].8'; 2025 '~Spare MB2[63].9'; 2026 '~Spare MB2[63].10'; 2027 '~S001CV1 - Conveyor Panel Disconnect Switch Not On MB2[63].11'; 2028 '~S001CV1Sfty- Conveyor Pull Cord #1 Tripped MB2[63].12'; 2029 '~S001CV1Sfty- Conveyor Pull Cord #2 Tripped MB2[63].13'; 2030 '~S001CV1Sfty- Conveyor Safety Contactor #1 (MC1) Still On MB2[63].14'; 2031 '~S001CV1Sfty- Conveyor Safety Contactor #1 (MC1) Not On MB2[63].15'; 2032 '~S001CV1Sfty- Conveyor Fwd Motor Starter (MF) Still On MB2[63].16'; 2033 '~S001CV1Sfty- Conveyor Fwd Motor Starter (MF) Not On MB2[63].17'; 2034 '~S001CV1Sfty- Conveyor Rev Motor Starter (MR) Still On MB2[63].18'; 2035 '~S001CV1Sfty- Conveyor Rev Motor Starter (MR) Not On MB2[63].19'; 2036 '~Spare MB2[63].20'; 2037 '~Spare MB2[63].21'; 2038 '~S001CV1 ~ Conveyor Auto/Mastering SS Not In Auto Postion MB2[63].22'; 2039 '~Spare MB2[63].23'; 2040 '~Spare MB2[63].24'; 2041 '~Spare MB2[63].25'; 2042 '~Spare MB2[63].26'; 2043 '~Spare MB2[63].27'; 2044 '~Spare MB2[63].28'; 2045 '~Spare MB2[63].29'; 2046 '~Spare MB2[63].30'; 2047 '~Spare MB2[63].31'; 2048 '~S003_004PRBDES1 - EtherNet Switch Connection Inhibited MB2[64].0'; 2049 '~Spare MB2[64].1'; 2050 '~Spare MB2[64].2'; 2051 '~S003_004PRBDV1 - Module Connection Inhibited MB2[64].3'; 2052 '~S003_004PRBDC - Module Connection Inhibited MB2[64].4'; 2053 '~S003_004PRB1B1 - Module Connection Inhibited MB2[64].5'; 2054 '~S003_004PRB1B2 - Module Connection Inhibited MB2[64].6'; 2055 '~Spare MB2[64].7'; 2056 '~Spare MB2[64].8'; 2057 '~Spare MB2[64].9'; 2058 '~S003_004PRB Panel Disconnect Off MB2[64].10'; 2059 '~S003PRB Motor Contactor 1MC Still On MB2[64].11'; 2060 '~S003PRB Motor Contactor 1MC Not On MB2[64].12'; 2061 '~S003PRB In Station Pallet/Skid Hold MB2[64].13'; 2062 '~Spare MB2[64].14'; 2063 '~S003PRB Motor Brake Relay 1BC1 Still On MB2[64].15'; 2064 '~S003PRB Motor Brake Relay 1BC1 Not On MB2[64].16'; 2065 '~S003PRB Motor Brake Relay 1BC2 Still On MB2[64].17'; 2066 '~S003PRB Motor Brake Relay 1BC2 Not On MB2[64].18'; 2067 '~S003Lft Lifter Contactor 1LMC Still On MB2[64].19'; 2068 '~S003Lft Lifter Contactor 1LMC Not On MB2[64].20'; 2069 '~Spare MB2[64].21'; 2070 '~S003LFT Lifter Safety Pin Fault MB2[64].22'; 2071 '~Spare MB2[64].23'; 2072 '~Spare MB2[64].24'; 2073 '~Spare MB2[64].25'; 2074 '~Spare MB2[64].26'; 2075 '~Spare MB2[64].27'; 2076 '~Spare MB2[64].28'; 2077 '~Spare MB2[64].29'; 2078 '~Spare MB2[64].30'; 2079 '~Spare MB2[64].31'; 2080 '~Spare MB2[65].0'; 2081 '~Spare MB2[65].1'; 2082 '~Spare MB2[65].2'; 2083 '~S003_004PRBDV2 - Module Connection Inhibited MB2[65].3'; 2084 '~Spare MB2[65].4'; 2085 '~S003_004PRB2B1 - Module Connection Inhibited MB2[65].5'; 2086 '~S003_004PRB2B2 - Module Connection Inhibited MB2[65].6'; 2087 '~Spare MB2[65].7'; 2088 '~Spare MB2[65].8'; 2089 '~Spare MB2[65].9'; 2090 '~Spare MB2[65].10'; 2091 '~S004PRB Motor Contactor 2MC Still On MB2[65].11'; 2092 '~S004PRB Motor Contactor 2MC Not On MB2[65].12'; 2093 '~S004PRB In Station Pallet/Skid 